// TIA Portal project "Automatizare_RT" (V17) (continued)
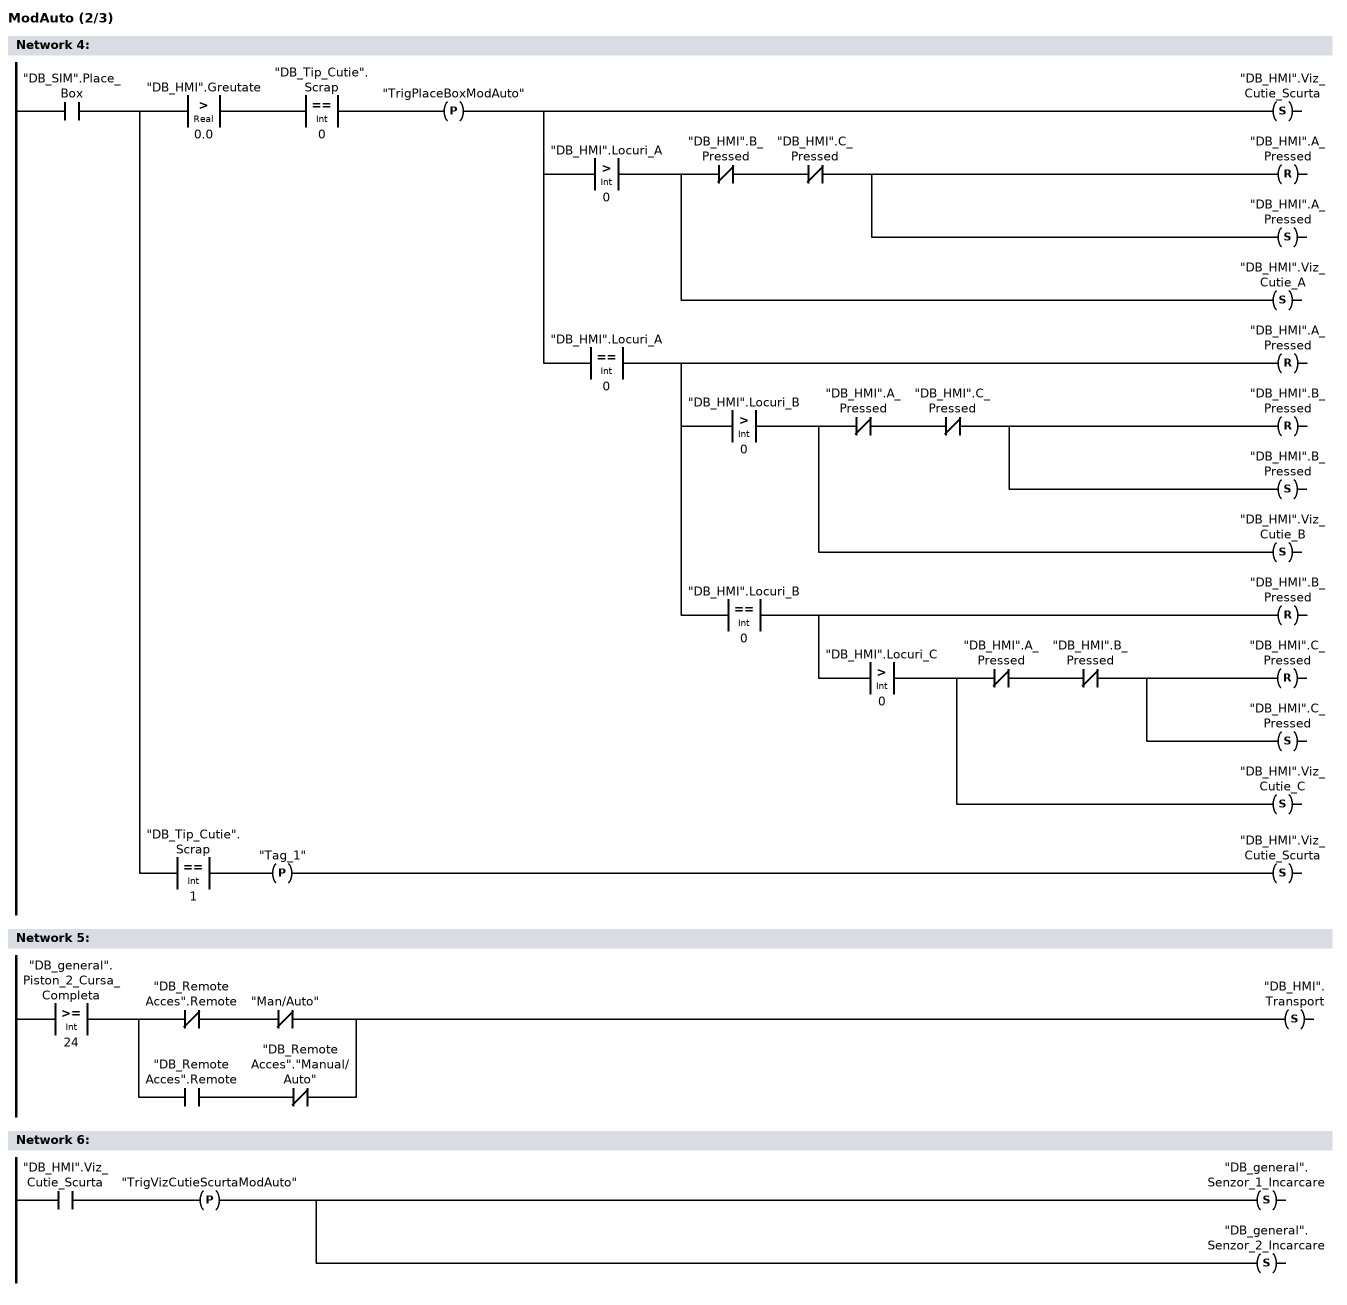
   RUNG wire#powerrail
      Contact( "DB_SIM".Place_Box )
      wire#w1
      { S7_Templates := "SrcType := Real" } GT_Contact(in1 := "DB_HMI".Greutate, in2 := 0.0)
      { S7_Templates := "SrcType := Int" } EQ_Contact(in1 := "DB_Tip_Cutie".Scrap, in2 := 0)
      P_Trig( "TrigPlaceBoxModAuto" )
      wire#w2
      S_Coil( "DB_HMI".Viz_Cutie_Scurta )
   END_RUNG
   RUNG wire#w2
      { S7_Templates := "SrcType := Int" } GT_Contact(in1 := "DB_HMI".Locuri_A, in2 := 0)
      wire#w3
      I_Contact( "DB_HMI".B_Pressed )
      I_Contact( "DB_HMI".C_Pressed )
      wire#w4
      R_Coil( "DB_HMI".A_Pressed )
   END_RUNG
   RUNG wire#w4
      S_Coil( "DB_HMI".A_Pressed )
   END_RUNG
   RUNG wire#w3
      S_Coil( "DB_HMI".Viz_Cutie_A )
   END_RUNG
   RUNG wire#w2
      { S7_Templates := "SrcType := Int" } EQ_Contact(in1 := "DB_HMI".Locuri_A, in2 := 0)
      wire#w5
      R_Coil( "DB_HMI".A_Pressed )
   END_RUNG
   RUNG wire#w5
      { S7_Templates := "SrcType := Int" } GT_Contact(in1 := "DB_HMI".Locuri_B, in2 := 0)
      wire#w6
      I_Contact( "DB_HMI".A_Pressed )
      I_Contact( "DB_HMI".C_Pressed )
      wire#w7
      R_Coil( "DB_HMI".B_Pressed )
   END_RUNG
   RUNG wire#w7
      S_Coil( "DB_HMI".B_Pressed )
   END_RUNG
   RUNG wire#w6
      S_Coil( "DB_HMI".Viz_Cutie_B )
   END_RUNG
   RUNG wire#w5
      { S7_Templates := "SrcType := Int" } EQ_Contact(in1 := "DB_HMI".Locuri_B, in2 := 0)
      wire#w8
      R_Coil( "DB_HMI".B_Pressed )
   END_RUNG
   RUNG wire#w8
      { S7_Templates := "SrcType := Int" } GT_Contact(in1 := "DB_HMI".Locuri_C, in2 := 0)
      wire#w9
      I_Contact( "DB_HMI".A_Pressed )
      I_Contact( "DB_HMI".B_Pressed )
      wire#w10
      R_Coil( "DB_HMI".C_Pressed )
   END_RUNG
   RUNG wire#w10
      S_Coil( "DB_HMI".C_Pressed )
   END_RUNG
   RUNG wire#w9
      S_Coil( "DB_HMI".Viz_Cutie_C )
   END_RUNG
   RUNG wire#w1
      { S7_Templates := "SrcType := Int" } EQ_Contact(in1 := "DB_Tip_Cutie".Scrap, in2 := 1)
      P_Trig( "Tag_1" )
      S_Coil( "DB_HMI".Viz_Cutie_Scurta )
   END_RUNG
   // the same network as SCL:
   #_w1 := "DB_SIM".Place_Box AND ("DB_HMI".Greutate > 0.0) AND ("DB_Tip_Cutie".Scrap = 0);
   #_w2 := #_w1 AND NOT "TrigPlaceBoxModAuto";   // rising edge
   "TrigPlaceBoxModAuto" := #_w1;
   IF #_w2 THEN "DB_HMI".Viz_Cutie_Scurta := TRUE; END_IF;
   #_w3 := #_w2 AND ("DB_HMI".Locuri_A > 0);
   IF #_w3 AND NOT "DB_HMI".B_Pressed AND NOT "DB_HMI".C_Pressed THEN
       "DB_HMI".A_Pressed := FALSE;
       "DB_HMI".A_Pressed := TRUE;
   END_IF;
   IF #_w3 THEN "DB_HMI".Viz_Cutie_A := TRUE; END_IF;
   #_w4 := #_w2 AND ("DB_HMI".Locuri_A = 0);
   IF #_w4 THEN "DB_HMI".A_Pressed := FALSE; END_IF;
   #_w5 := #_w4 AND ("DB_HMI".Locuri_B > 0);
   IF #_w5 AND NOT "DB_HMI".A_Pressed AND NOT "DB_HMI".C_Pressed THEN
       "DB_HMI".B_Pressed := FALSE;
       "DB_HMI".B_Pressed := TRUE;
   END_IF;
   IF #_w5 THEN "DB_HMI".Viz_Cutie_B := TRUE; END_IF;
   #_w6 := #_w4 AND ("DB_HMI".Locuri_B = 0);
   IF #_w6 THEN "DB_HMI".B_Pressed := FALSE; END_IF;
   #_w7 := #_w6 AND ("DB_HMI".Locuri_C > 0);
   IF #_w7 AND NOT "DB_HMI".A_Pressed AND NOT "DB_HMI".B_Pressed THEN
       "DB_HMI".C_Pressed := FALSE;
       "DB_HMI".C_Pressed := TRUE;
   END_IF;
   IF #_w7 THEN "DB_HMI".Viz_Cutie_C := TRUE; END_IF;
   #_w8 := "DB_SIM".Place_Box AND ("DB_Tip_Cutie".Scrap = 1);
   #_w9 := #_w8 AND NOT "Tag_1";   // rising edge
   "Tag_1" := #_w8;
   IF #_w9 THEN "DB_HMI".Viz_Cutie_Scurta := TRUE; END_IF;
END_REGION

REGION Network 5
   RUNG wire#powerrail
      { S7_Templates := "SrcType := Int" } GE_Contact(in1 := "DB_general".Piston_2_Cursa_Completa, in2 := 24)
      wire#w1
      I_Contact( "DB_RemoteAcces".Remote )
      I_Contact( "Man/Auto" )
      wire#w2
      S_Coil( "DB_HMI".Transport )
   END_RUNG
   RUNG wire#w1
      Contact( "DB_RemoteAcces".Remote )
      I_Contact( "DB_RemoteAcces"."Manual/Auto" )
   END_RUNG wire#w2
   // the same network as SCL:
   IF ("DB_general".Piston_2_Cursa_Completa >= 24) AND ((NOT "DB_RemoteAcces".Remote AND NOT "Man/Auto") OR ("DB_RemoteAcces".Remote AND NOT "DB_RemoteAcces"."Manual/Auto")) THEN
       "DB_HMI".Transport := TRUE;
   END_IF;
END_REGION

REGION Network 6
   RUNG wire#powerrail
      Contact( "DB_HMI".Viz_Cutie_Scurta )
      P_Trig( "TrigVizCutieScurtaModAuto" )
      wire#w1
      S_Coil( "DB_general".Senzor_1_Incarcare )
   END_RUNG
   RUNG wire#w1
      S_Coil( "DB_general".Senzor_2_Incarcare )
   END_RUNG
   // the same network as SCL:
   #_w1 := "DB_HMI".Viz_Cutie_Scurta AND NOT "TrigVizCutieScurtaModAuto";   // rising edge
   "TrigVizCutieScurtaModAuto" := "DB_HMI".Viz_Cutie_Scurta;
   IF #_w1 THEN
       "DB_general".Senzor_1_Incarcare := TRUE;
       "DB_general".Senzor_2_Incarcare := TRUE;
   END_IF;
END_REGION

REGION Network 7
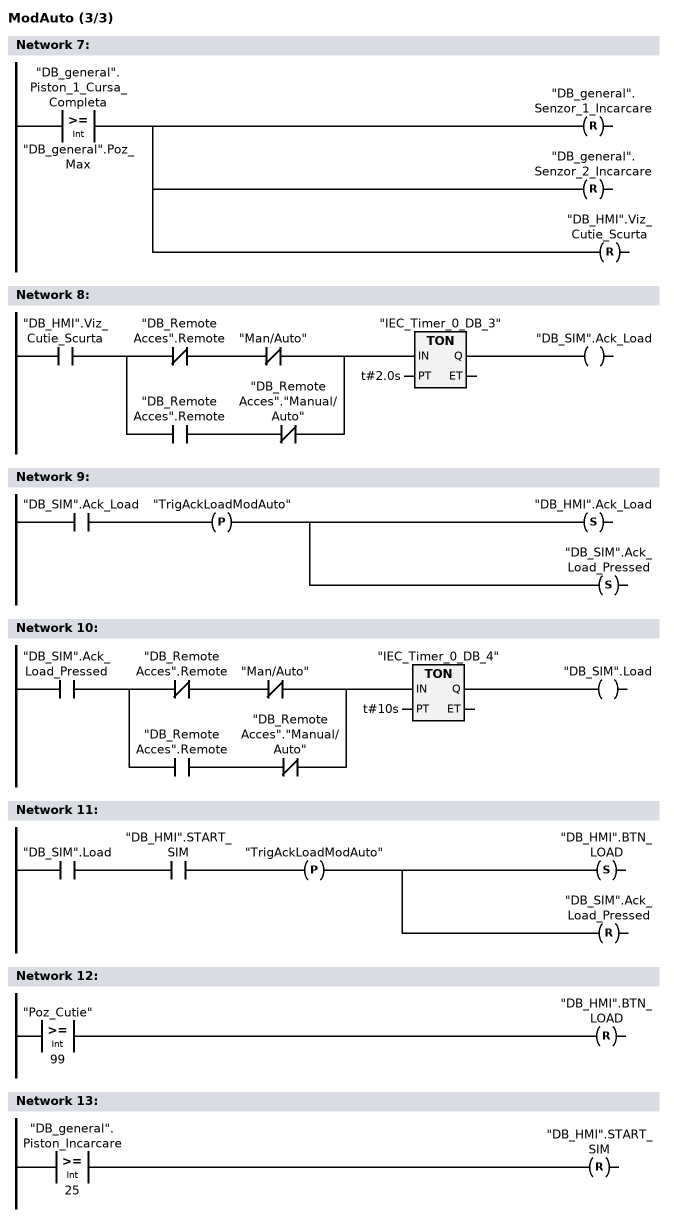
   RUNG wire#powerrail
      { S7_Templates := "SrcType := Int" } GE_Contact(in1 := "DB_general".Piston_1_Cursa_Completa, in2 := "DB_general".Poz_Max)
      wire#w1
      R_Coil( "DB_general".Senzor_1_Incarcare )
   END_RUNG
   RUNG wire#w1
      R_Coil( "DB_general".Senzor_2_Incarcare )
   END_RUNG
   RUNG wire#w1
      R_Coil( "DB_HMI".Viz_Cutie_Scurta )
   END_RUNG
   // the same network as SCL:
   IF "DB_general".Piston_1_Cursa_Completa >= "DB_general".Poz_Max THEN
       "DB_general".Senzor_1_Incarcare := FALSE;
       "DB_general".Senzor_2_Incarcare := FALSE;
       "DB_HMI".Viz_Cutie_Scurta := FALSE;
   END_IF;
END_REGION

REGION Network 8
   "IEC_Timer_0_DB_3".TON(IN := "DB_HMI".Viz_Cutie_Scurta AND ((NOT "DB_RemoteAcces".Remote AND NOT "Man/Auto") OR ("DB_RemoteAcces".Remote AND NOT "DB_RemoteAcces"."Manual/Auto")),
                          PT := t#2.0s);
   "DB_SIM".Ack_Load := "IEC_Timer_0_DB_3".Q;
END_REGION

REGION Network 9
   RUNG wire#powerrail
      Contact( "DB_SIM".Ack_Load )
      P_Trig( "TrigAckLoadModAuto" )
      wire#w1
      S_Coil( "DB_HMI".Ack_Load )
   END_RUNG
   RUNG wire#w1
      S_Coil( "DB_SIM".Ack_Load_Pressed )
   END_RUNG
   // the same network as SCL:
   #_w1 := "DB_SIM".Ack_Load AND NOT "TrigAckLoadModAuto";   // rising edge
   "TrigAckLoadModAuto" := "DB_SIM".Ack_Load;
   IF #_w1 THEN
       "DB_HMI".Ack_Load := TRUE;
       "DB_SIM".Ack_Load_Pressed := TRUE;
   END_IF;
END_REGION

REGION Network 10
   "IEC_Timer_0_DB_4".TON(IN := "DB_SIM".Ack_Load_Pressed AND ((NOT "DB_RemoteAcces".Remote AND NOT "Man/Auto") OR ("DB_RemoteAcces".Remote AND NOT "DB_RemoteAcces"."Manual/Auto")),
                          PT := t#10s);
   "DB_SIM".Load := "IEC_Timer_0_DB_4".Q;
END_REGION

REGION Network 11
   RUNG wire#powerrail
      Contact( "DB_SIM".Load )
      Contact( "DB_HMI".START_SIM )
      P_Trig( "TrigAckLoadModAuto" )
      wire#w1
      S_Coil( "DB_HMI".BTN_LOAD )
   END_RUNG
   RUNG wire#w1
      R_Coil( "DB_SIM".Ack_Load_Pressed )
   END_RUNG
   // the same network as SCL:
   #_w1 := "DB_SIM".Load AND "DB_HMI".START_SIM;
   #_w2 := #_w1 AND NOT "TrigAckLoadModAuto";   // rising edge
   "TrigAckLoadModAuto" := #_w1;
   IF #_w2 THEN
       "DB_HMI".BTN_LOAD := TRUE;
       "DB_SIM".Ack_Load_Pressed := FALSE;
   END_IF;
END_REGION

REGION Network 12
   RUNG wire#powerrail
      { S7_Templates := "SrcType := Int" } GE_Contact(in1 := "Poz_Cutie", in2 := 99)
      R_Coil( "DB_HMI".BTN_LOAD )
   END_RUNG
   // the same network as SCL:
   IF "Poz_Cutie" >= 99 THEN "DB_HMI".BTN_LOAD := FALSE; END_IF;
END_REGION

REGION Network 13
   RUNG wire#powerrail
      { S7_Templates := "SrcType := Int" } GE_Contact(in1 := "DB_general".Piston_Incarcare, in2 := 25)
      R_Coil( "DB_HMI".START_SIM )
   END_RUNG
   // the same network as SCL:
   IF "DB_general".Piston_Incarcare >= 25 THEN "DB_HMI".START_SIM := FALSE; END_IF;
END_REGION
END_FUNCTION_BLOCK

FUNCTION "Emg_Stop_Fcn" : Void   // FC4, LAD
{ S7_Optimized_Access := 'FALSE' }
VERSION : 0.1
BEGIN

REGION Network 1
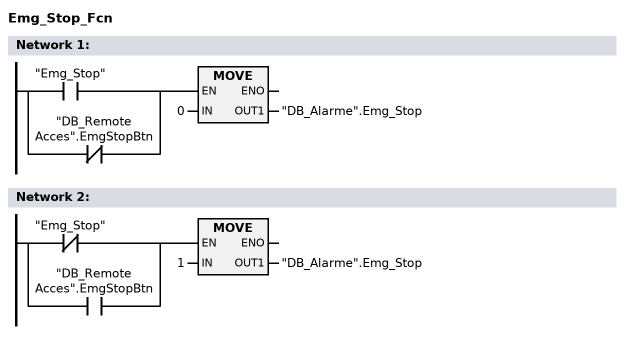
   RUNG wire#powerrail
      Contact( "Emg_Stop" )
      wire#w1
      { S7_GenerateENO := "TRUE" } Move(in := 0, out1 => "DB_Alarme".Emg_Stop)
   END_RUNG
   RUNG wire#powerrail
      I_Contact( "DB_RemoteAcces".EmgStopBtn )
   END_RUNG wire#w1
   // the same network as SCL:
   IF "Emg_Stop" OR NOT "DB_RemoteAcces".EmgStopBtn THEN "DB_Alarme".Emg_Stop := 0; END_IF;
END_REGION

REGION Network 2
   RUNG wire#powerrail
      I_Contact( "Emg_Stop" )
      wire#w1
      { S7_GenerateENO := "TRUE" } Move(in := 1, out1 => "DB_Alarme".Emg_Stop)
   END_RUNG
   RUNG wire#powerrail
      Contact( "DB_RemoteAcces".EmgStopBtn )
   END_RUNG wire#w1
   // the same network as SCL:
   IF NOT "Emg_Stop" OR "DB_RemoteAcces".EmgStopBtn THEN "DB_Alarme".Emg_Stop := 1; END_IF;
END_REGION
END_FUNCTION

FUNCTION "Vizibilitate_Manuale/Automate" : Void   // FC5, STL
{ S7_Optimized_Access := 'FALSE' }
VERSION : 0.1
BEGIN

REGION Network 1
         A     "DB_HMI".Viz_Cutie_Banda_1;
         A(;
         L     "DB_HMI".Tip_Cutie_Lung;
         L     1;
         ==I;
         );
         JNB   Label_0;
         L     1;
         T     "DB_HMI"."Viz_Cutie_Man/Auto";
   Label_0:NOP   0;
END_REGION

REGION Network 2
         A     "DB_HMI".Viz_Cutie_Banda_1;
         A(;
         L     "DB_HMI".Tip_Cutie_Lung;
         L     2;
         ==I;
         );
         JNB   Label_1;
         L     2;
         T     "DB_HMI"."Viz_Cutie_Man/Auto";
   Label_1:NOP   0;
END_REGION

REGION Network 3
         AN    "DB_HMI".Viz_Cutie_Banda_1;
         JNB   Label_2;
         L     0;
         T     "DB_HMI"."Viz_Cutie_Man/Auto";
   Label_2:NOP   0;
END_REGION

REGION Network 4
         A     "DB_HMI".Viz_Cutie_Scurta;
         A(;
         L     "DB_HMI".Tip_Cutie_Lung;
         L     1;
         ==I;
         );
         JNB   Label_3;
         L     1;
         T     "DB_Tranzitii"."Tip_Cutie_Man/Auto_Start";
   Label_3:NOP   0;
END_REGION

REGION Network 5
         A     "DB_HMI".Viz_Cutie_Scurta;
         A(;
         L     "DB_HMI".Tip_Cutie_Lung;
         L     2;
         ==I;
         );
         JNB   Label_4;
         L     2;
         T     "DB_Tranzitii"."Tip_Cutie_Man/Auto_Start";
   Label_4:NOP   0;
END_REGION

REGION Network 6
         A(;
         O(;
         L     "DB_general".Piston_1_Cursa_Completa;
         L     25;
         ==I;
         );
         ON    "DB_HMI".Viz_Cutie_Scurta;
         );
         JNB   Label_5;
         L     0;
         T     "DB_Tranzitii"."Tip_Cutie_Man/Auto_Start";
   Label_5:NOP   0;
END_REGION

REGION Network 7
         A(;
         L     "Poz_Cutie";
         L     99;
         ==I;
         );
         A(;
         L     "DB_HMI".Tip_Cutie_Lung;
         L     1;
         ==I;
         );
         FP    "TrigVizCutiePoz99CutieLung1";
         JNB   Label_6;
         L     1;
         T     "DB_Tranzitii"."TipCutieMan/Auto_End";
   Label_6:NOP   0;
END_REGION

REGION Network 8
         A(;
         L     "Poz_Cutie";
         L     99;
         ==I;
         );
         A(;
         L     "DB_HMI".Tip_Cutie_Lung;
         L     2;
         ==I;
         );
         FP    "TrigPozCutie99CutieLung2";
         JNB   Label_7;
         L     2;
         T     "DB_Tranzitii"."TipCutieMan/Auto_End";
   Label_7:NOP   0;
END_REGION

REGION Network 9
         A(;
         O(;
         L     "Poz_Cutie";
         L     99;
         <I;
         );
         O(;
         L     "DB_general".Piston_2_Cursa_Completa;
         L     20;
         >I;
         );
         );
         JNB   Label_8;
         L     0;
         T     "DB_Tranzitii"."TipCutieMan/Auto_End";
   Label_8:NOP   0;
END_REGION
END_FUNCTION

FUNCTION "Status_Pistoane" : Void   // FC7, LAD
{ S7_Optimized_Access := 'FALSE' }
VERSION : 0.1
BEGIN

REGION Network 1: Cand Piston1 este in functiune / Wenn Kolben 1 in Betrieb ist
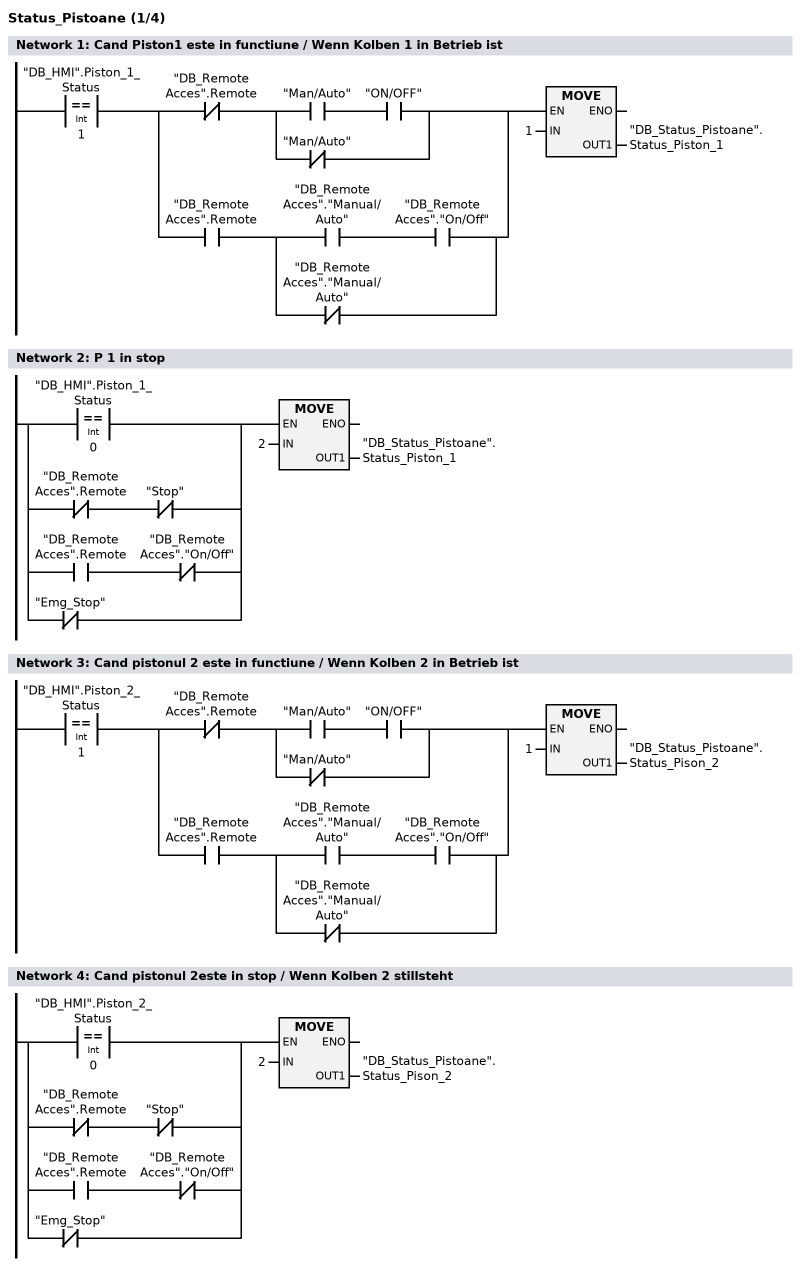
   RUNG wire#powerrail
      { S7_Templates := "SrcType := Int" } EQ_Contact(in1 := "DB_HMI".Piston_1_Status, in2 := 1)
      wire#w1
      I_Contact( "DB_RemoteAcces".Remote )
      wire#w2
      Contact( "Man/Auto" )
      Contact( "ON/OFF" )
      wire#w3
      { S7_GenerateENO := "TRUE" } Move(in := 1, out1 => "DB_Status_Pistoane".Status_Piston_1)
   END_RUNG
   RUNG wire#w2
      I_Contact( "Man/Auto" )
   END_RUNG wire#w3
   RUNG wire#w1
      Contact( "DB_RemoteAcces".Remote )
      wire#w4
      Contact( "DB_RemoteAcces"."Manual/Auto" )
      Contact( "DB_RemoteAcces"."On/Off" )
   END_RUNG wire#w3
   RUNG wire#w4
      I_Contact( "DB_RemoteAcces"."Manual/Auto" )
   END_RUNG wire#w3
   // the same network as SCL:
   IF ("DB_HMI".Piston_1_Status = 1) AND ((NOT "DB_RemoteAcces".Remote AND (("Man/Auto" AND "ON/OFF") OR NOT "Man/Auto")) OR ("DB_RemoteAcces".Remote AND (("DB_RemoteAcces"."Manual/Auto" AND "DB_RemoteAcces"."On/Off") OR NOT "DB_RemoteAcces"."Manual/Auto"))) THEN
       "DB_Status_Pistoane".Status_Piston_1 := 1;
   END_IF;
END_REGION

REGION Network 2: P 1 in stop
   RUNG wire#powerrail
      { S7_Templates := "SrcType := Int" } EQ_Contact(in1 := "DB_HMI".Piston_1_Status, in2 := 0)
      wire#w1
      { S7_GenerateENO := "TRUE" } Move(in := 2, out1 => "DB_Status_Pistoane".Status_Piston_1)
   END_RUNG
   RUNG wire#powerrail
      I_Contact( "DB_RemoteAcces".Remote )
      I_Contact( "Stop" )
   END_RUNG wire#w1
   RUNG wire#powerrail
      Contact( "DB_RemoteAcces".Remote )
      I_Contact( "DB_RemoteAcces"."On/Off" )
   END_RUNG wire#w1
   RUNG wire#powerrail
      I_Contact( "Emg_Stop" )
   END_RUNG wire#w1
   // the same network as SCL:
   IF ("DB_HMI".Piston_1_Status = 0) OR (NOT "DB_RemoteAcces".Remote AND NOT "Stop") OR ("DB_RemoteAcces".Remote AND NOT "DB_RemoteAcces"."On/Off") OR NOT "Emg_Stop" THEN
       "DB_Status_Pistoane".Status_Piston_1 := 2;
   END_IF;
END_REGION

REGION Network 3: Cand pistonul 2 este in functiune / Wenn Kolben 2 in Betrieb ist
   RUNG wire#powerrail
      { S7_Templates := "SrcType := Int" } EQ_Contact(in1 := "DB_HMI".Piston_2_Status, in2 := 1)
      wire#w1
      I_Contact( "DB_RemoteAcces".Remote )
      wire#w2
      Contact( "Man/Auto" )
      Contact( "ON/OFF" )
      wire#w3
      { S7_GenerateENO := "TRUE" } Move(in := 1, out1 => "DB_Status_Pistoane".Status_Pison_2)
   END_RUNG
   RUNG wire#w2
      I_Contact( "Man/Auto" )
   END_RUNG wire#w3
   RUNG wire#w1
      Contact( "DB_RemoteAcces".Remote )
      wire#w4
      Contact( "DB_RemoteAcces"."Manual/Auto" )
      Contact( "DB_RemoteAcces"."On/Off" )
   END_RUNG wire#w3
   RUNG wire#w4
      I_Contact( "DB_RemoteAcces"."Manual/Auto" )
   END_RUNG wire#w3
   // the same network as SCL:
   IF ("DB_HMI".Piston_2_Status = 1) AND ((NOT "DB_RemoteAcces".Remote AND (("Man/Auto" AND "ON/OFF") OR NOT "Man/Auto")) OR ("DB_RemoteAcces".Remote AND (("DB_RemoteAcces"."Manual/Auto" AND "DB_RemoteAcces"."On/Off") OR NOT "DB_RemoteAcces"."Manual/Auto"))) THEN
       "DB_Status_Pistoane".Status_Pison_2 := 1;
   END_IF;
END_REGION

REGION Network 4: Cand pistonul 2este in stop / Wenn Kolben 2 stillsteht
   RUNG wire#powerrail
      { S7_Templates := "SrcType := Int" } EQ_Contact(in1 := "DB_HMI".Piston_2_Status, in2 := 0)
      wire#w1
      { S7_GenerateENO := "TRUE" } Move(in := 2, out1 => "DB_Status_Pistoane".Status_Pison_2)
   END_RUNG
   RUNG wire#powerrail
      I_Contact( "DB_RemoteAcces".Remote )
      I_Contact( "Stop" )
   END_RUNG wire#w1
   RUNG wire#powerrail
      Contact( "DB_RemoteAcces".Remote )
      I_Contact( "DB_RemoteAcces"."On/Off" )
   END_RUNG wire#w1
   RUNG wire#powerrail
      I_Contact( "Emg_Stop" )
   END_RUNG wire#w1
   // the same network as SCL:
   IF ("DB_HMI".Piston_2_Status = 0) OR (NOT "DB_RemoteAcces".Remote AND NOT "Stop") OR ("DB_RemoteAcces".Remote AND NOT "DB_RemoteAcces"."On/Off") OR NOT "Emg_Stop" THEN
       "DB_Status_Pistoane".Status_Pison_2 := 2;
   END_IF;
END_REGION

REGION Network 5: Piston A este in functiune / Kolben A ist in Betrieb
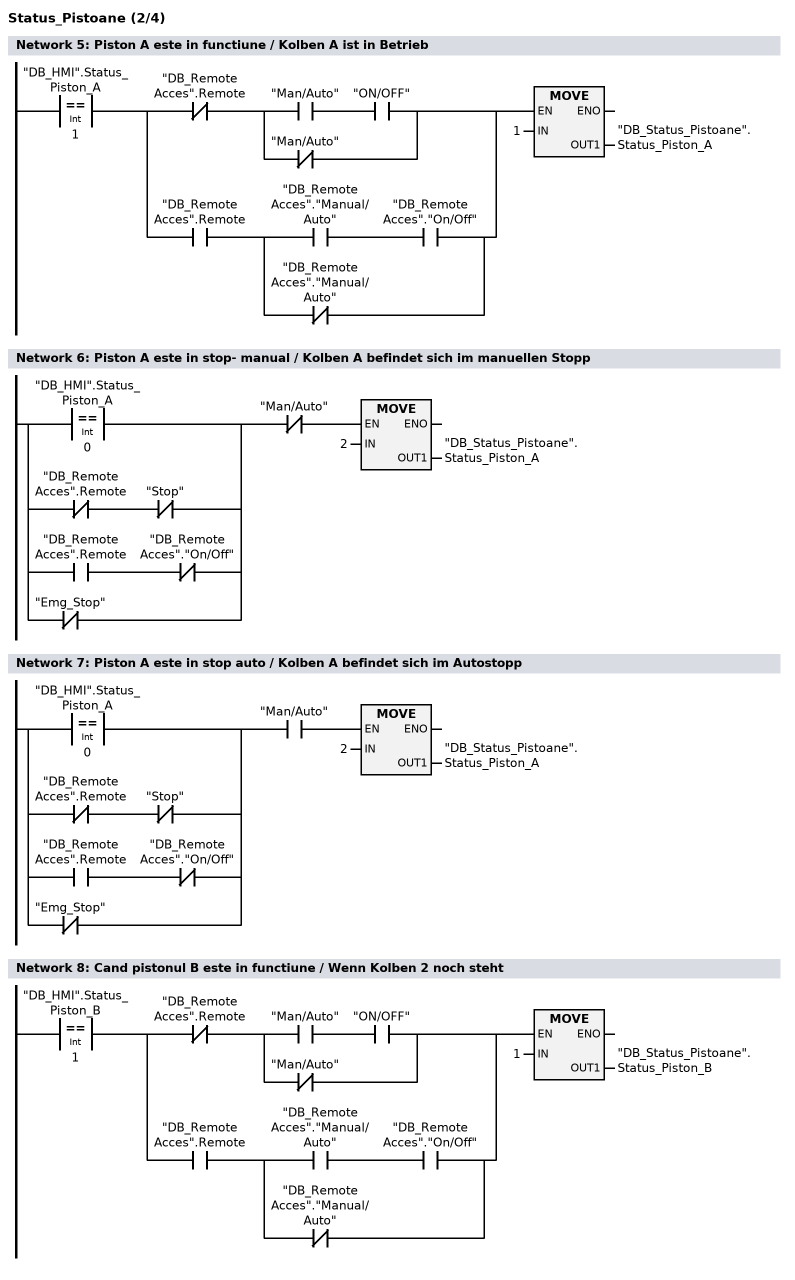
   RUNG wire#powerrail
      { S7_Templates := "SrcType := Int" } EQ_Contact(in1 := "DB_HMI".Status_Piston_A, in2 := 1)
      wire#w1
      I_Contact( "DB_RemoteAcces".Remote )
      wire#w2
      Contact( "Man/Auto" )
      Contact( "ON/OFF" )
      wire#w3
      { S7_GenerateENO := "TRUE" } Move(in := 1, out1 => "DB_Status_Pistoane".Status_Piston_A)
   END_RUNG
   RUNG wire#w2
      I_Contact( "Man/Auto" )
   END_RUNG wire#w3
   RUNG wire#w1
      Contact( "DB_RemoteAcces".Remote )
      wire#w4
      Contact( "DB_RemoteAcces"."Manual/Auto" )
      Contact( "DB_RemoteAcces"."On/Off" )
   END_RUNG wire#w3
   RUNG wire#w4
      I_Contact( "DB_RemoteAcces"."Manual/Auto" )
   END_RUNG wire#w3
   // the same network as SCL:
   IF ("DB_HMI".Status_Piston_A = 1) AND ((NOT "DB_RemoteAcces".Remote AND (("Man/Auto" AND "ON/OFF") OR NOT "Man/Auto")) OR ("DB_RemoteAcces".Remote AND (("DB_RemoteAcces"."Manual/Auto" AND "DB_RemoteAcces"."On/Off") OR NOT "DB_RemoteAcces"."Manual/Auto"))) THEN
       "DB_Status_Pistoane".Status_Piston_A := 1;
   END_IF;
END_REGION

REGION Network 6: Piston A este in stop- manual / Kolben A befindet sich im manuellen Stopp
   RUNG wire#powerrail
      { S7_Templates := "SrcType := Int" } EQ_Contact(in1 := "DB_HMI".Status_Piston_A, in2 := 0)
      wire#w1
      I_Contact( "Man/Auto" )
      { S7_GenerateENO := "TRUE" } Move(in := 2, out1 => "DB_Status_Pistoane".Status_Piston_A)
   END_RUNG
   RUNG wire#powerrail
      I_Contact( "DB_RemoteAcces".Remote )
      I_Contact( "Stop" )
   END_RUNG wire#w1
   RUNG wire#powerrail
      Contact( "DB_RemoteAcces".Remote )
      I_Contact( "DB_RemoteAcces"."On/Off" )
   END_RUNG wire#w1
   RUNG wire#powerrail
      I_Contact( "Emg_Stop" )
   END_RUNG wire#w1
   // the same network as SCL:
   IF (("DB_HMI".Status_Piston_A = 0) OR (NOT "DB_RemoteAcces".Remote AND NOT "Stop") OR ("DB_RemoteAcces".Remote AND NOT "DB_RemoteAcces"."On/Off") OR NOT "Emg_Stop") AND NOT "Man/Auto" THEN
       "DB_Status_Pistoane".Status_Piston_A := 2;
   END_IF;
END_REGION

REGION Network 7: Piston A este in stop auto / Kolben A befindet sich im Autostopp
   RUNG wire#powerrail
      { S7_Templates := "SrcType := Int" } EQ_Contact(in1 := "DB_HMI".Status_Piston_A, in2 := 0)
      wire#w1
      Contact( "Man/Auto" )
      { S7_GenerateENO := "TRUE" } Move(in := 2, out1 => "DB_Status_Pistoane".Status_Piston_A)
   END_RUNG
   RUNG wire#powerrail
      I_Contact( "DB_RemoteAcces".Remote )
      I_Contact( "Stop" )
   END_RUNG wire#w1
   RUNG wire#powerrail
      Contact( "DB_RemoteAcces".Remote )
      I_Contact( "DB_RemoteAcces"."On/Off" )
   END_RUNG wire#w1
   RUNG wire#powerrail
      I_Contact( "Emg_Stop" )
   END_RUNG wire#w1
   // the same network as SCL:
   IF (("DB_HMI".Status_Piston_A = 0) OR (NOT "DB_RemoteAcces".Remote AND NOT "Stop") OR ("DB_RemoteAcces".Remote AND NOT "DB_RemoteAcces"."On/Off") OR NOT "Emg_Stop") AND "Man/Auto" THEN
       "DB_Status_Pistoane".Status_Piston_A := 2;
   END_IF;
END_REGION

REGION Network 8: Cand pistonul B este in functiune / Wenn Kolben 2 noch steht
   RUNG wire#powerrail
      { S7_Templates := "SrcType := Int" } EQ_Contact(in1 := "DB_HMI".Status_Piston_B, in2 := 1)
      wire#w1
      I_Contact( "DB_RemoteAcces".Remote )
      wire#w2
      Contact( "Man/Auto" )
      Contact( "ON/OFF" )
      wire#w3
      { S7_GenerateENO := "TRUE" } Move(in := 1, out1 => "DB_Status_Pistoane".Status_Piston_B)
   END_RUNG
   RUNG wire#w2
      I_Contact( "Man/Auto" )
   END_RUNG wire#w3
   RUNG wire#w1
      Contact( "DB_RemoteAcces".Remote )
      wire#w4
      Contact( "DB_RemoteAcces"."Manual/Auto" )
      Contact( "DB_RemoteAcces"."On/Off" )
   END_RUNG wire#w3
   RUNG wire#w4
      I_Contact( "DB_RemoteAcces"."Manual/Auto" )
   END_RUNG wire#w3
   // the same network as SCL:
   IF ("DB_HMI".Status_Piston_B = 1) AND ((NOT "DB_RemoteAcces".Remote AND (("Man/Auto" AND "ON/OFF") OR NOT "Man/Auto")) OR ("DB_RemoteAcces".Remote AND (("DB_RemoteAcces"."Manual/Auto" AND "DB_RemoteAcces"."On/Off") OR NOT "DB_RemoteAcces"."Manual/Auto"))) THEN
       "DB_Status_Pistoane".Status_Piston_B := 1;
   END_IF;
END_REGION

REGION Network 9: Piston B este in stop- manual / Kolben B befindet sich im manuellen Stopp
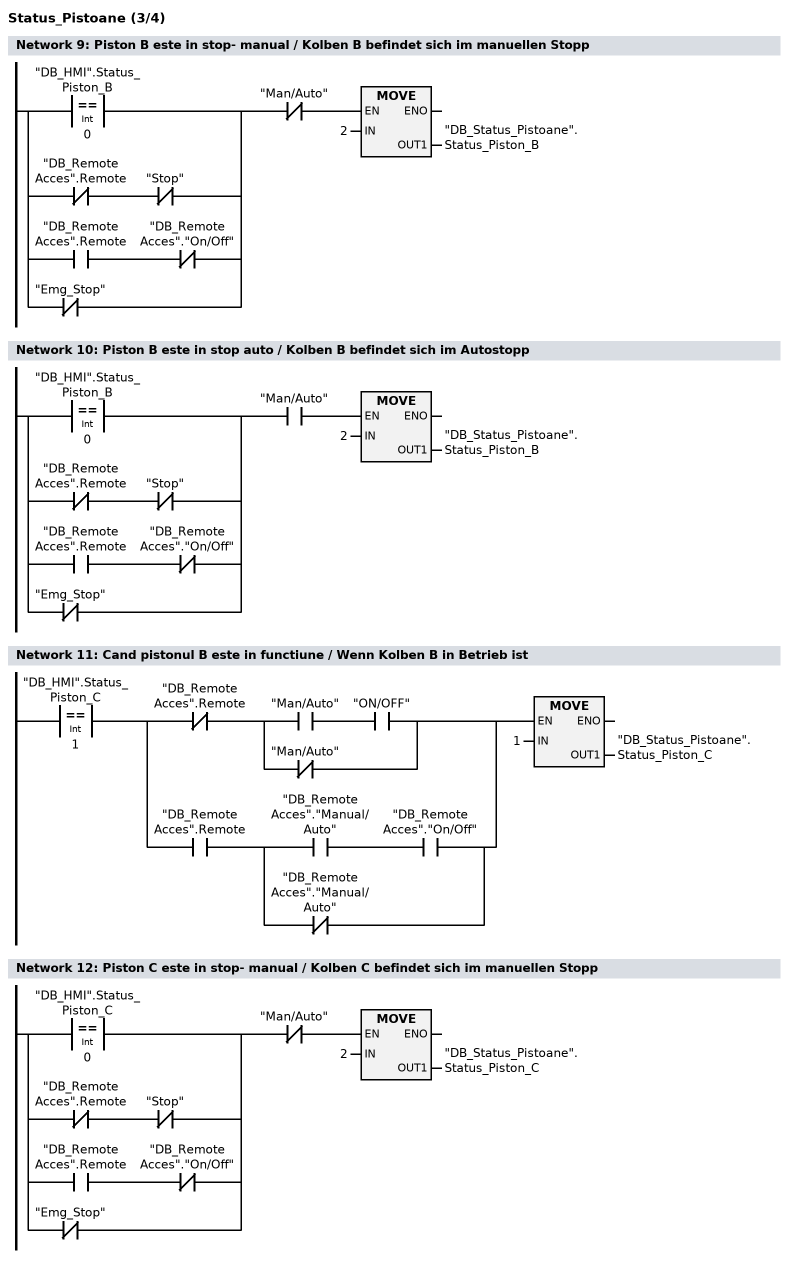
   RUNG wire#powerrail
      { S7_Templates := "SrcType := Int" } EQ_Contact(in1 := "DB_HMI".Status_Piston_B, in2 := 0)
      wire#w1
      I_Contact( "Man/Auto" )
      { S7_GenerateENO := "TRUE" } Move(in := 2, out1 => "DB_Status_Pistoane".Status_Piston_B)
   END_RUNG
   RUNG wire#powerrail
      I_Contact( "DB_RemoteAcces".Remote )
      I_Contact( "Stop" )
   END_RUNG wire#w1
   RUNG wire#powerrail
      Contact( "DB_RemoteAcces".Remote )
      I_Contact( "DB_RemoteAcces"."On/Off" )
   END_RUNG wire#w1
   RUNG wire#powerrail
      I_Contact( "Emg_Stop" )
   END_RUNG wire#w1
   // the same network as SCL:
   IF (("DB_HMI".Status_Piston_B = 0) OR (NOT "DB_RemoteAcces".Remote AND NOT "Stop") OR ("DB_RemoteAcces".Remote AND NOT "DB_RemoteAcces"."On/Off") OR NOT "Emg_Stop") AND NOT "Man/Auto" THEN
       "DB_Status_Pistoane".Status_Piston_B := 2;
   END_IF;
END_REGION

REGION Network 10: Piston B este in stop auto / Kolben B befindet sich im Autostopp
   RUNG wire#powerrail
      { S7_Templates := "SrcType := Int" } EQ_Contact(in1 := "DB_HMI".Status_Piston_B, in2 := 0)
      wire#w1
      Contact( "Man/Auto" )
      { S7_GenerateENO := "TRUE" } Move(in := 2, out1 => "DB_Status_Pistoane".Status_Piston_B)
   END_RUNG
   RUNG wire#powerrail
      I_Contact( "DB_RemoteAcces".Remote )
      I_Contact( "Stop" )
   END_RUNG wire#w1
   RUNG wire#powerrail
      Contact( "DB_RemoteAcces".Remote )
      I_Contact( "DB_RemoteAcces"."On/Off" )
   END_RUNG wire#w1
   RUNG wire#powerrail
      I_Contact( "Emg_Stop" )
   END_RUNG wire#w1
   // the same network as SCL:
   IF (("DB_HMI".Status_Piston_B = 0) OR (NOT "DB_RemoteAcces".Remote AND NOT "Stop") OR ("DB_RemoteAcces".Remote AND NOT "DB_RemoteAcces"."On/Off") OR NOT "Emg_Stop") AND "Man/Auto" THEN
       "DB_Status_Pistoane".Status_Piston_B := 2;
   END_IF;
END_REGION

REGION Network 11: Cand pistonul B este in functiune / Wenn Kolben B in Betrieb ist
   RUNG wire#powerrail
      { S7_Templates := "SrcType := Int" } EQ_Contact(in1 := "DB_HMI".Status_Piston_C, in2 := 1)
      wire#w1
      I_Contact( "DB_RemoteAcces".Remote )
      wire#w2
      Contact( "Man/Auto" )
      Contact( "ON/OFF" )
      wire#w3
      { S7_GenerateENO := "TRUE" } Move(in := 1, out1 => "DB_Status_Pistoane".Status_Piston_C)
   END_RUNG
   RUNG wire#w2
      I_Contact( "Man/Auto" )
   END_RUNG wire#w3
   RUNG wire#w1
      Contact( "DB_RemoteAcces".Remote )
      wire#w4
      Contact( "DB_RemoteAcces"."Manual/Auto" )
      Contact( "DB_RemoteAcces"."On/Off" )
   END_RUNG wire#w3
   RUNG wire#w4
      I_Contact( "DB_RemoteAcces"."Manual/Auto" )
   END_RUNG wire#w3
   // the same network as SCL:
   IF ("DB_HMI".Status_Piston_C = 1) AND ((NOT "DB_RemoteAcces".Remote AND (("Man/Auto" AND "ON/OFF") OR NOT "Man/Auto")) OR ("DB_RemoteAcces".Remote AND (("DB_RemoteAcces"."Manual/Auto" AND "DB_RemoteAcces"."On/Off") OR NOT "DB_RemoteAcces"."Manual/Auto"))) THEN
       "DB_Status_Pistoane".Status_Piston_C := 1;
   END_IF;
END_REGION

REGION Network 12: Piston C este in stop- manual / Kolben C befindet sich im manuellen Stopp
   RUNG wire#powerrail
      { S7_Templates := "SrcType := Int" } EQ_Contact(in1 := "DB_HMI".Status_Piston_C, in2 := 0)
      wire#w1
      I_Contact( "Man/Auto" )
      { S7_GenerateENO := "TRUE" } Move(in := 2, out1 => "DB_Status_Pistoane".Status_Piston_C)
   END_RUNG
   RUNG wire#powerrail
      I_Contact( "DB_RemoteAcces".Remote )
      I_Contact( "Stop" )
   END_RUNG wire#w1
   RUNG wire#powerrail
      Contact( "DB_RemoteAcces".Remote )
      I_Contact( "DB_RemoteAcces"."On/Off" )
   END_RUNG wire#w1
   RUNG wire#powerrail
      I_Contact( "Emg_Stop" )
   END_RUNG wire#w1
   // the same network as SCL:
   IF (("DB_HMI".Status_Piston_C = 0) OR (NOT "DB_RemoteAcces".Remote AND NOT "Stop") OR ("DB_RemoteAcces".Remote AND NOT "DB_RemoteAcces"."On/Off") OR NOT "Emg_Stop") AND NOT "Man/Auto" THEN
       "DB_Status_Pistoane".Status_Piston_C := 2;
   END_IF;
END_REGION

REGION Network 13: Piston C este in stop auto / Kolben C befindet sich im Autostopp
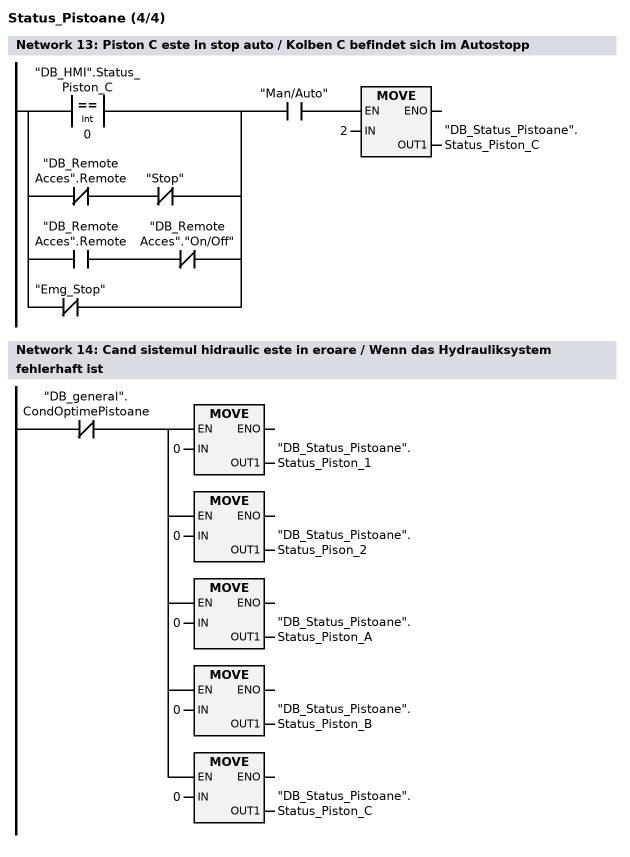
   RUNG wire#powerrail
      { S7_Templates := "SrcType := Int" } EQ_Contact(in1 := "DB_HMI".Status_Piston_C, in2 := 0)
      wire#w1
      Contact( "Man/Auto" )
      { S7_GenerateENO := "TRUE" } Move(in := 2, out1 => "DB_Status_Pistoane".Status_Piston_C)
   END_RUNG
   RUNG wire#powerrail
      I_Contact( "DB_RemoteAcces".Remote )
      I_Contact( "Stop" )
   END_RUNG wire#w1
   RUNG wire#powerrail
      Contact( "DB_RemoteAcces".Remote )
      I_Contact( "DB_RemoteAcces"."On/Off" )
   END_RUNG wire#w1
   RUNG wire#powerrail
      I_Contact( "Emg_Stop" )
   END_RUNG wire#w1
   // the same network as SCL:
   IF (("DB_HMI".Status_Piston_C = 0) OR (NOT "DB_RemoteAcces".Remote AND NOT "Stop") OR ("DB_RemoteAcces".Remote AND NOT "DB_RemoteAcces"."On/Off") OR NOT "Emg_Stop") AND "Man/Auto" THEN
       "DB_Status_Pistoane".Status_Piston_C := 2;
   END_IF;
END_REGION
